REGION Network 7 (SCL): Head #4
   "M256_Manag_IDB".M256F_IDB[3].INPUT_xPressureDec :="i.1B414AP1.1B414SA1.Head4.CuttingPressure-";
   "M256_Manag_IDB".M256A_IDB[3].INPUT_xCarriageInWorkPosition := "i.1B414AP1.1B414SQ1.Head4.CarriageHeadWorkPosition";
   "M256_Manag_IDB".M256F_IDB[3].INPUT_xPressureInc := "i.1B414AP1.1B414SA1.Head4.CuttingPressure+";
   "Z256".INPUT_rgxHeadsInProduction[3] := "i.1B414AP1.1B414SA2.Head4.ProductionON";
   "M256_Manag_IDB".M256F_IDB[3].INPUT_xForceFiring := 0;
   "M256_Manag_IDB".M256A_IDB[3].INPUT_xForceArming := 0;
   "M256_Manag_IDB".M256M_IDB[3].INPUT_xBrakeRelease := FALSE;
   "M256_Manag_IDB".M256M_IDB[3].INPUT_xOverstroke := TRUE;//"i.1B410AP1.1B291KA4.Head4-5.CarriageTraslationAntiCollision";
END_REGION

REGION Network 8 (SCL): Head #5
   "M256_Manag_IDB".M256F_IDB[4].INPUT_xPressureDec := "i.1B415AP1.1B415SA1.Head5.CuttingPressure-";
   "M256_Manag_IDB".M256A_IDB[4].INPUT_xCarriageInWorkPosition := "i.1B415AP1.1B415SQ1.Head5.CarriageHeadWorkPosition";
   "M256_Manag_IDB".M256F_IDB[4].INPUT_xPressureInc := "i.1B415AP1.1B415SA1.Head5.CuttingPressure+";
   "Z256".INPUT_rgxHeadsInProduction[4] :="i.1B415AP1.1B415SA2.Head5.ProductionON";
   "M256_Manag_IDB".M256F_IDB[4].INPUT_xForceFiring := 0;
   "M256_Manag_IDB".M256A_IDB[4].INPUT_xForceArming := 0;
   "M256_Manag_IDB".M256M_IDB[4].INPUT_xBrakeRelease := FALSE;
   "M256_Manag_IDB".M256M_IDB[4].INPUT_xOverstroke := TRUE;//"i.1B410AP1.1B291KA5.Head5-6.CarriageTraslationAntiCollision";
END_REGION

REGION Network 9 (SCL): Head #6 / Head #5
   "M256_Manag_IDB".M256F_IDB[5].INPUT_xPressureDec := "i.1B416AP1.1B416SA1.Head6.CuttingPressure-";
   "M256_Manag_IDB".M256A_IDB[5].INPUT_xCarriageInWorkPosition := "i.1B416AP1.1B416SQ1.Head6.CarriageHeadWorkPosition";
   "M256_Manag_IDB".M256F_IDB[5].INPUT_xPressureInc := "i.1B416AP1.1B416SA1.Head6.CuttingPressure+";
   "Z256".INPUT_rgxHeadsInProduction[5] :="i.1B416AP1.1B416SA2.Head6.ProductionON";
   "M256_Manag_IDB".M256F_IDB[5].INPUT_xForceFiring := 0;
   "M256_Manag_IDB".M256A_IDB[5].INPUT_xForceArming := 0;
   "M256_Manag_IDB".M256M_IDB[5].INPUT_xBrakeRelease := FALSE;
   "M256_Manag_IDB".M256M_IDB[5].INPUT_xOverstroke := TRUE;//"i.1B410AP1.1B291KA8.Head6-7.CarriageTraslationAntiCollision";
END_REGION

REGION Network 10 (SCL): Head #7 / Head #5
   "M256_Manag_IDB".M256F_IDB[6].INPUT_xPressureDec := "i.1B417AP1.1B417SA1.Head7.CuttingPressure-";
   "M256_Manag_IDB".M256A_IDB[6].INPUT_xCarriageInWorkPosition := "i.1B417AP1.1B417SQ1.Head7.CarriageHeadWorkPosition";
   "M256_Manag_IDB".M256F_IDB[6].INPUT_xPressureInc := "i.1B417AP1.1B417SA1.Head7.CuttingPressure+";
   "Z256".INPUT_rgxHeadsInProduction[6] :="i.1B417AP1.1B417SA2.Head7.ProductionON";
   "M256_Manag_IDB".M256F_IDB[6].INPUT_xForceFiring := 0;
   "M256_Manag_IDB".M256A_IDB[6].INPUT_xForceArming := 0;
   "M256_Manag_IDB".M256M_IDB[6].INPUT_xBrakeRelease := FALSE;
   "M256_Manag_IDB".M256M_IDB[6].INPUT_xOverstroke := TRUE;//"i.1B410AP1.1B291KA7.Head7-8.CarriageTraslationAntiCollision";
END_REGION

REGION Network 11 (SCL): Head #8 / Head #5
   "M256_Manag_IDB".M256F_IDB[7].INPUT_xPressureDec := "i.1B418AP1.1B418SA1.Head8.CuttingPressure-";
   "M256_Manag_IDB".M256A_IDB[7].INPUT_xCarriageInWorkPosition := "i.1B418AP1.1B418SQ1.Head8.CarriageHeadWorkPosition";
   "M256_Manag_IDB".M256F_IDB[7].INPUT_xPressureInc := "i.1B418AP1.1B418SA1.Head8.CuttingPressure+";
   "Z256".INPUT_rgxHeadsInProduction[7] :="i.1B418AP1.1B418SA2.Head8.ProductionON";
   "M256_Manag_IDB".M256F_IDB[7].INPUT_xForceFiring := 0;
   "M256_Manag_IDB".M256A_IDB[7].INPUT_xForceArming := 0;
   "M256_Manag_IDB".M256M_IDB[7].INPUT_xBrakeRelease := FALSE;
   "M256_Manag_IDB".M256M_IDB[7].INPUT_xOverstroke := TRUE;//"i.1B410AP1.1B291KA8.Head8-9.CarriageTraslationAntiCollision";
END_REGION

REGION Network 12 (SCL): IDevice
   "CM_IDEV_FromMainLine" := "i.IDeviceCPU0";
END_REGION
END_FUNCTION

FUNCTION "M256M_SbrCheckCollision" : Void   // FC10, SCL
{ S7_Optimized_Access := 'TRUE' }
VERSION : 0.1
   VAR_OUTPUT
      o_rgxHeadVirtualCollision : Array[0.."CONST_dNumberOfHeadsCycle"] of Bool;
   END_VAR
   VAR_TEMP
      TMP_dIndex : DInt;
      TMP_xCollision : Bool;
      TMP_xCollisionNext : Bool;
      TMP_dActHeadPosition_cmm : DInt;
      TMP_dNextHeadPosition_cmm : DInt;
   END_VAR
BEGIN
   ////--------------------------------------------------------------------------------------------------------------------
   //   Copyright (c)  Bottero Spa
   //--------------------------------------------------------------
   //   Routine: NomeRoutine
   //       Author: Alberto Cigliutti
   //   Created: July 2016
   //--------------------------------------------------------------
   //   Description: This routine will analize the data out from the manager, and compile 
   //  a collision array
   //
   //   History:
   //
   ////--------------------------------------------------------------------------------------------------------------------

   FOR #TMP_dIndex := 0 TO "CONST_dNumberOfHeadsCycle" DO
       #o_rgxHeadVirtualCollision[#TMP_dIndex] := 0;
   END_FOR;

   FOR #TMP_dIndex := 0 TO "CONST_dNumberOfHeadsCycle" DO

       #TMP_xCollision := 0;
       #TMP_xCollisionNext := 0;

       IF #TMP_dIndex = 0 OR #TMP_dIndex = "CONST_dNumberOfHeadsCycle" THEN
           //For the first head and last head, we check the position request, if is less then the home
           //we rise a virtual collision
           IF NOT "PLANT_CONSTANTS".CONST_rgxHomeSide[#TMP_dIndex] AND
               ("Z256_Manager".tOutputData.rgdHeadsPositions_cmm[#TMP_dIndex] < "M256_Manag_IDB".M256M_IDB[#TMP_dIndex].tHMR.dHeadHomePositions_cmm) THEN

               #TMP_xCollision := 1;
               #o_rgxHeadVirtualCollision[#TMP_dIndex] := #TMP_xCollision;

           ELSIF ("PLANT_CONSTANTS".CONST_rgxHomeSide[#TMP_dIndex] AND
               "Z256_Manager".tOutputData.rgdHeadsPositions_cmm[#TMP_dIndex]>"M256_Manag_IDB".M256M_IDB[#TMP_dIndex].tHMR.dHeadHomePositions_cmm) THEN

               #TMP_xCollision := 1;
               #o_rgxHeadVirtualCollision[#TMP_dIndex] := #TMP_xCollision;
           END_IF;
       END_IF;

       //Start to search the next head position,
       //only jump this check on the last head
       IF #TMP_dIndex < "CONST_dNumberOfHeadsCycle" THEN

           #TMP_dActHeadPosition_cmm := "Z256_Manager".tOutputData.rgdHeadsPositions_cmm[#TMP_dIndex] + "PLANT_CONSTANTS".CONST_dHOppoSideEnc_cmm[#TMP_dIndex];
           #TMP_dNextHeadPosition_cmm := "Z256_Manager".tOutputData.rgdHeadsPositions_cmm[#TMP_dIndex + 1] - "PLANT_CONSTANTS".CONST_dHOpSideEnc_cmm[#TMP_dIndex + 1];

           IF (#TMP_dActHeadPosition_cmm > #TMP_dNextHeadPosition_cmm) THEN
               #TMP_xCollision := 1;
               #TMP_xCollisionNext := 1;
           END_IF;

           #o_rgxHeadVirtualCollision[#TMP_dIndex + 1] := #TMP_xCollisionNext;
           #o_rgxHeadVirtualCollision[#TMP_dIndex] := #TMP_xCollision;

       END_IF;



   END_FOR;
END_FUNCTION

FUNCTION "M256M_HMI_Logics" : Void   // FC11, LAD
{ S7_Optimized_Access := 'TRUE' }
VERSION : 0.1
   VAR_IN_OUT
      io_ST_xHeadReferredSwitch : Array[0.."CONST_dNumberOfHeadsCycle"] of Bool;
   END_VAR
   VAR_TEMP
      TMP_dIndex : DInt;
   END_VAR
   VAR_TEMP   // added for the SCL form of the ladder/FBD networks
      _w1 : Bool;
   END_VAR
BEGIN

REGION Network 1: #####_HMI_LOGICS_#####
END_REGION

REGION Network 2 (SCL): Force heads homing
   IF "Z256_hmi".tHMW.xForceHeadsHoming THEN
       FOR #TMP_dIndex := 0 TO "CONST_dNumberOfHeadsCycle" DO
           #io_ST_xHeadReferredSwitch[#TMP_dIndex] := 0;
       END_FOR;
       "Z256_hmi".tHMW.xForceHeadsHoming := false;
   END_IF;
END_REGION

REGION Network 3: Calibration function allowed
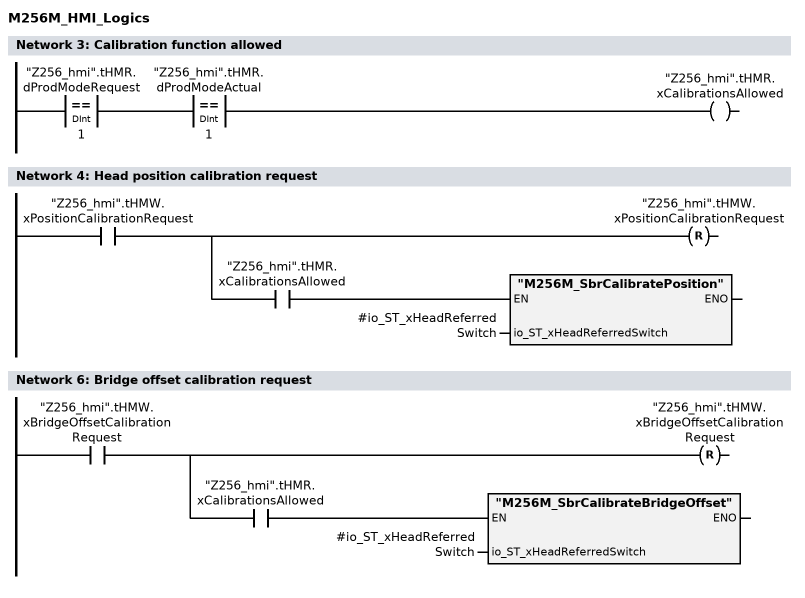
   RUNG wire#powerrail
      { S7_Templates := "SrcType := DInt" } EQ_Contact(in1 := "Z256_hmi".tHMR.dProdModeRequest, in2 := 1)
      { S7_Templates := "SrcType := DInt" } EQ_Contact(in1 := "Z256_hmi".tHMR.dProdModeActual, in2 := 1)
      Coil( "Z256_hmi".tHMR.xCalibrationsAllowed )
   END_RUNG
   // the same network as SCL:
   "Z256_hmi".tHMR.xCalibrationsAllowed := ("Z256_hmi".tHMR.dProdModeRequest = 1) AND ("Z256_hmi".tHMR.dProdModeActual = 1);
END_REGION

REGION Network 4: Head position calibration request
   RUNG wire#powerrail
      Contact( "Z256_hmi".tHMW.xPositionCalibrationRequest )
      wire#w1
      R_Coil( "Z256_hmi".tHMW.xPositionCalibrationRequest )
   END_RUNG
   RUNG wire#w1
      Contact( "Z256_hmi".tHMR.xCalibrationsAllowed )
      "M256M_SbrCalibratePosition"(io_ST_xHeadReferredSwitch := #io_ST_xHeadReferredSwitch)
   END_RUNG
   // the same network as SCL:
   #_w1 := "Z256_hmi".tHMW.xPositionCalibrationRequest;
   IF #_w1 THEN "Z256_hmi".tHMW.xPositionCalibrationRequest := FALSE; END_IF;
   IF #_w1 AND "Z256_hmi".tHMR.xCalibrationsAllowed THEN
       "M256M_SbrCalibratePosition"(io_ST_xHeadReferredSwitch := #io_ST_xHeadReferredSwitch);
   END_IF;
END_REGION

REGION Network 5 (SCL): Update home head
   FOR #TMP_dIndex := 0 TO "CONST_dNumberOfHeadsCycle" DO
       IF "M256_Manag_IDB".M256M_IDB[#TMP_dIndex].tHMW.xUpdateHomeHead THEN
           "M256_Manag_IDB".M256M_IDB[#TMP_dIndex].tHMW.xUpdateHomeHead := 0; 
           "M256_Manag_IDB".M256M_IDB[#TMP_dIndex].tHMR.dHeadHomePositions_cmm := "M256_Manag_IDB".M256M_IDB[#TMP_dIndex].tHMW.dHeadHomePositions_cmm;
       END_IF;
   END_FOR;
END_REGION

REGION Network 6: Bridge offset calibration request
   RUNG wire#powerrail
      Contact( "Z256_hmi".tHMW.xBridgeOffsetCalibrationRequest )
      wire#w1
      R_Coil( "Z256_hmi".tHMW.xBridgeOffsetCalibrationRequest )
   END_RUNG
   RUNG wire#w1
      Contact( "Z256_hmi".tHMR.xCalibrationsAllowed )
      "M256M_SbrCalibrateBridgeOffset"(io_ST_xHeadReferredSwitch := #io_ST_xHeadReferredSwitch)
   END_RUNG
   // the same network as SCL:
   #_w1 := "Z256_hmi".tHMW.xBridgeOffsetCalibrationRequest;
   IF #_w1 THEN "Z256_hmi".tHMW.xBridgeOffsetCalibrationRequest := FALSE; END_IF;
   IF #_w1 AND "Z256_hmi".tHMR.xCalibrationsAllowed THEN
       "M256M_SbrCalibrateBridgeOffset"(io_ST_xHeadReferredSwitch := #io_ST_xHeadReferredSwitch);
   END_IF;
END_REGION
END_FUNCTION

FUNCTION "Encoder_Manager" : Void   // FC12, LAD
{ S7_Optimized_Access := 'TRUE' }
VERSION : 0.1
   VAR_TEMP
      TMP_rDummy : Real;
      TMP_dDummy : DInt;
      TMP_dIndex : DInt;
   END_VAR
   VAR_TEMP   // added for the SCL form of the ladder/FBD networks
      _w1 : Bool;
   END_VAR
BEGIN

REGION Network 1: Enable card counter
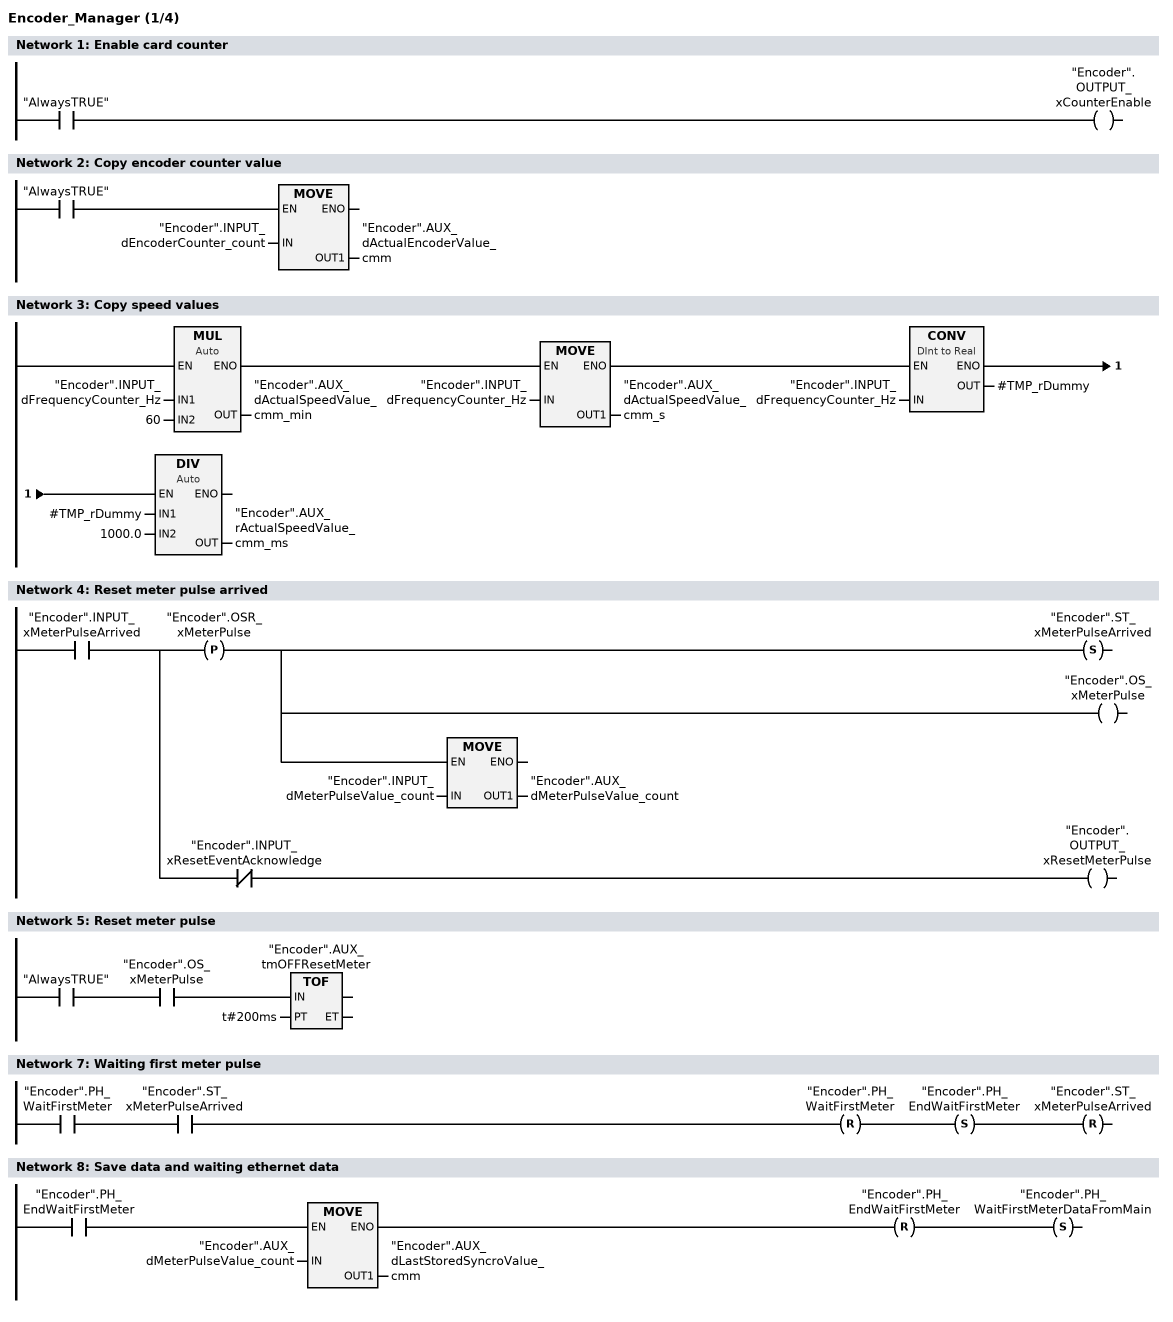
   RUNG wire#powerrail
      Contact( "AlwaysTRUE" )
      Coil( "Encoder".OUTPUT_xCounterEnable )
   END_RUNG
   // the same network as SCL:
   "Encoder".OUTPUT_xCounterEnable := "AlwaysTRUE";
END_REGION

REGION Network 2: Copy encoder counter value
   RUNG wire#powerrail
      Contact( "AlwaysTRUE" )
      Move(in := "Encoder".INPUT_dEncoderCounter_count, out1 => "Encoder".AUX_dActualEncoderValue_cmm)
   END_RUNG
   // the same network as SCL:
   IF "AlwaysTRUE" THEN
       "Encoder".AUX_dActualEncoderValue_cmm := "Encoder".INPUT_dEncoderCounter_count;
   END_IF;
END_REGION

REGION Network 3: Copy speed values
   RUNG wire#powerrail
      Mul(in1 := "Encoder".INPUT_dFrequencyCounter_Hz, in2 := 60, out => "Encoder".AUX_dActualSpeedValue_cmm_min)
      Move(in := "Encoder".INPUT_dFrequencyCounter_Hz, out1 => "Encoder".AUX_dActualSpeedValue_cmm_s)
      { S7_Templates := "[SrcType := DInt, DestType := Real]" } Convert(in := "Encoder".INPUT_dFrequencyCounter_Hz, out => #TMP_rDummy)
      Div(in1 := #TMP_rDummy, in2 := 1000.0, out => "Encoder".AUX_rActualSpeedValue_cmm_ms)
   END_RUNG
   // the same network as SCL:
   "Encoder".AUX_dActualSpeedValue_cmm_min := "Encoder".INPUT_dFrequencyCounter_Hz * 60;
   "Encoder".AUX_dActualSpeedValue_cmm_s := "Encoder".INPUT_dFrequencyCounter_Hz;
   #TMP_rDummy := DINT_TO_REAL("Encoder".INPUT_dFrequencyCounter_Hz);
   "Encoder".AUX_rActualSpeedValue_cmm_ms := #TMP_rDummy / 1000.0;
END_REGION

REGION Network 4: Reset meter pulse arrived
   RUNG wire#powerrail
      Contact( "Encoder".INPUT_xMeterPulseArrived )
      wire#w1
      P_Trig( "Encoder".OSR_xMeterPulse )
      wire#w2
      S_Coil( "Encoder".ST_xMeterPulseArrived )
   END_RUNG
   RUNG wire#w2
      Coil( "Encoder".OS_xMeterPulse )
   END_RUNG
   RUNG wire#w2
      Move(in := "Encoder".INPUT_dMeterPulseValue_count, out1 => "Encoder".AUX_dMeterPulseValue_count)
   END_RUNG
   RUNG wire#w1
      I_Contact( "Encoder".INPUT_xResetEventAcknowledge )
      Coil( "Encoder".OUTPUT_xResetMeterPulse )
   END_RUNG
   // the same network as SCL:
   #_w1 := "Encoder".INPUT_xMeterPulseArrived AND NOT "Encoder".OSR_xMeterPulse;   // rising edge
   "Encoder".OSR_xMeterPulse := "Encoder".INPUT_xMeterPulseArrived;
   IF #_w1 THEN "Encoder".ST_xMeterPulseArrived := TRUE; END_IF;
   "Encoder".OS_xMeterPulse := #_w1;
   IF #_w1 THEN "Encoder".AUX_dMeterPulseValue_count := "Encoder".INPUT_dMeterPulseValue_count; END_IF;
   "Encoder".OUTPUT_xResetMeterPulse := "Encoder".INPUT_xMeterPulseArrived AND NOT "Encoder".INPUT_xResetEventAcknowledge;
END_REGION

REGION Network 5: Reset meter pulse
   "Encoder".AUX_tmOFFResetMeter.TOF(IN := "AlwaysTRUE" AND "Encoder".OS_xMeterPulse, PT := t#200ms);
END_REGION

REGION Network 6: ### FIRST METER PHASES ###
END_REGION

REGION Network 7: Waiting first meter pulse
   RUNG wire#powerrail
      Contact( "Encoder".PH_WaitFirstMeter )
      Contact( "Encoder".ST_xMeterPulseArrived )
      R_Coil( "Encoder".PH_WaitFirstMeter )
      S_Coil( "Encoder".PH_EndWaitFirstMeter )
      R_Coil( "Encoder".ST_xMeterPulseArrived )
   END_RUNG
   // the same network as SCL:
   #_w1 := "Encoder".PH_WaitFirstMeter AND "Encoder".ST_xMeterPulseArrived;
   IF #_w1 THEN
       "Encoder".PH_WaitFirstMeter := FALSE;
       "Encoder".PH_EndWaitFirstMeter := TRUE;
       "Encoder".ST_xMeterPulseArrived := FALSE;
   END_IF;
END_REGION

REGION Network 8: Save data and waiting ethernet data
   RUNG wire#powerrail
      Contact( "Encoder".PH_EndWaitFirstMeter )
      Move(in := "Encoder".AUX_dMeterPulseValue_count, out1 => "Encoder".AUX_dLastStoredSyncroValue_cmm)
      R_Coil( "Encoder".PH_EndWaitFirstMeter )
      S_Coil( "Encoder".PH_WaitFirstMeterDataFromMain )
   END_RUNG
   // the same network as SCL:
   IF "Encoder".PH_EndWaitFirstMeter THEN
       "Encoder".AUX_dLastStoredSyncroValue_cmm := "Encoder".AUX_dMeterPulseValue_count;
   END_IF;
   #_w1 := "Encoder".PH_EndWaitFirstMeter;
   IF #_w1 THEN
       "Encoder".PH_EndWaitFirstMeter := FALSE;
       "Encoder".PH_WaitFirstMeterDataFromMain := TRUE;
   END_IF;
END_REGION

REGION Network 9: End waiting ethernet data
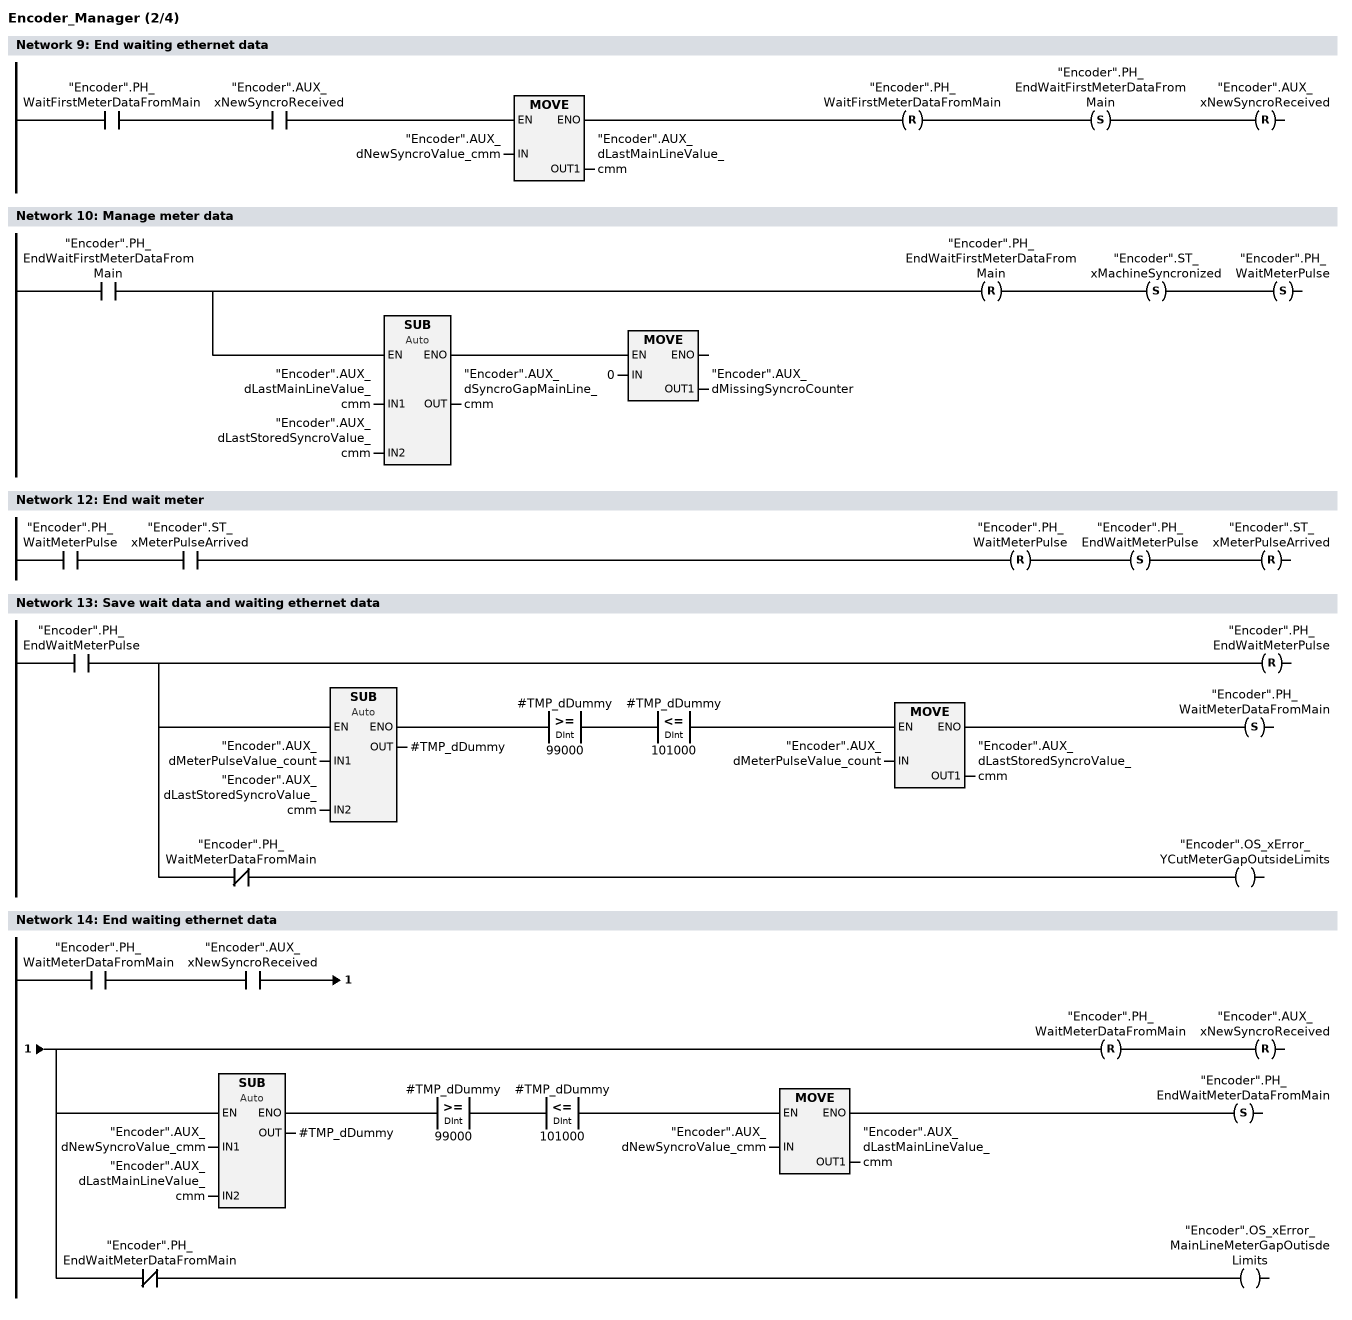
   RUNG wire#powerrail
      Contact( "Encoder".PH_WaitFirstMeterDataFromMain )
      Contact( "Encoder".AUX_xNewSyncroReceived )
      Move(in := "Encoder".AUX_dNewSyncroValue_cmm, out1 => "Encoder".AUX_dLastMainLineValue_cmm)
      R_Coil( "Encoder".PH_WaitFirstMeterDataFromMain )
      S_Coil( "Encoder".PH_EndWaitFirstMeterDataFromMain )
      R_Coil( "Encoder".AUX_xNewSyncroReceived )
   END_RUNG
   // the same network as SCL:
   IF "Encoder".PH_WaitFirstMeterDataFromMain AND "Encoder".AUX_xNewSyncroReceived THEN
       "Encoder".AUX_dLastMainLineValue_cmm := "Encoder".AUX_dNewSyncroValue_cmm;
   END_IF;
   #_w1 := "Encoder".PH_WaitFirstMeterDataFromMain AND "Encoder".AUX_xNewSyncroReceived;
   IF #_w1 THEN
       "Encoder".PH_WaitFirstMeterDataFromMain := FALSE;
       "Encoder".PH_EndWaitFirstMeterDataFromMain := TRUE;
       "Encoder".AUX_xNewSyncroReceived := FALSE;
   END_IF;
END_REGION

REGION Network 10: Manage meter data
   RUNG wire#powerrail
      Contact( "Encoder".PH_EndWaitFirstMeterDataFromMain )
      wire#w1
      R_Coil( "Encoder".PH_EndWaitFirstMeterDataFromMain )
      S_Coil( "Encoder".ST_xMachineSyncronized )
      S_Coil( "Encoder".PH_WaitMeterPulse )
   END_RUNG
   RUNG wire#w1
      Sub(in1 := "Encoder".AUX_dLastMainLineValue_cmm, in2 := "Encoder".AUX_dLastStoredSyncroValue_cmm, out => "Encoder".AUX_dSyncroGapMainLine_cmm)
      Move(in := 0, out1 => "Encoder".AUX_dMissingSyncroCounter)
   END_RUNG
   // the same network as SCL:
   #_w1 := "Encoder".PH_EndWaitFirstMeterDataFromMain;
   IF #_w1 THEN
       "Encoder".PH_EndWaitFirstMeterDataFromMain := FALSE;
       "Encoder".ST_xMachineSyncronized := TRUE;
       "Encoder".PH_WaitMeterPulse := TRUE;
       "Encoder".AUX_dSyncroGapMainLine_cmm := "Encoder".AUX_dLastMainLineValue_cmm - "Encoder".AUX_dLastStoredSyncroValue_cmm;
       "Encoder".AUX_dMissingSyncroCounter := 0;
   END_IF;
END_REGION

REGION Network 11: ### METER PHASES ###
END_REGION

REGION Network 12: End wait meter
   RUNG wire#powerrail
      Contact( "Encoder".PH_WaitMeterPulse )
      Contact( "Encoder".ST_xMeterPulseArrived )
      R_Coil( "Encoder".PH_WaitMeterPulse )
      S_Coil( "Encoder".PH_EndWaitMeterPulse )
      R_Coil( "Encoder".ST_xMeterPulseArrived )
   END_RUNG
   // the same network as SCL:
   #_w1 := "Encoder".PH_WaitMeterPulse AND "Encoder".ST_xMeterPulseArrived;
   IF #_w1 THEN
       "Encoder".PH_WaitMeterPulse := FALSE;
       "Encoder".PH_EndWaitMeterPulse := TRUE;
       "Encoder".ST_xMeterPulseArrived := FALSE;
   END_IF;
END_REGION

REGION Network 13: Save wait data and waiting ethernet data
   RUNG wire#powerrail
      Contact( "Encoder".PH_EndWaitMeterPulse )
      wire#w1
      R_Coil( "Encoder".PH_EndWaitMeterPulse )
   END_RUNG
   RUNG wire#w1
      Sub(in1 := "Encoder".AUX_dMeterPulseValue_count, in2 := "Encoder".AUX_dLastStoredSyncroValue_cmm, out => #TMP_dDummy)
      { S7_Templates := "SrcType := DInt" } GE_Contact(in1 := #TMP_dDummy, in2 := 99000)
      { S7_Templates := "SrcType := DInt" } LE_Contact(in1 := #TMP_dDummy, in2 := 101000)
      Move(in := "Encoder".AUX_dMeterPulseValue_count, out1 => "Encoder".AUX_dLastStoredSyncroValue_cmm)
      S_Coil( "Encoder".PH_WaitMeterDataFromMain )
   END_RUNG
   RUNG wire#w1
      I_Contact( "Encoder".PH_WaitMeterDataFromMain )
      Coil( "Encoder".OS_xError_YCutMeterGapOutsideLimits )
   END_RUNG
   // the same network as SCL:
   #_w1 := "Encoder".PH_EndWaitMeterPulse;
   IF #_w1 THEN
       "Encoder".PH_EndWaitMeterPulse := FALSE;
       #TMP_dDummy := "Encoder".AUX_dMeterPulseValue_count - "Encoder".AUX_dLastStoredSyncroValue_cmm;
   END_IF;
   IF #_w1 AND (#TMP_dDummy >= 99000) AND (#TMP_dDummy <= 101000) THEN
       "Encoder".AUX_dLastStoredSyncroValue_cmm := "Encoder".AUX_dMeterPulseValue_count;
       "Encoder".PH_WaitMeterDataFromMain := TRUE;
   END_IF;
   "Encoder".OS_xError_YCutMeterGapOutsideLimits := #_w1 AND NOT "Encoder".PH_WaitMeterDataFromMain;
END_REGION

REGION Network 14: End waiting ethernet data
   RUNG wire#powerrail
      Contact( "Encoder".PH_WaitMeterDataFromMain )
      Contact( "Encoder".AUX_xNewSyncroReceived )
      wire#w1
      R_Coil( "Encoder".PH_WaitMeterDataFromMain )
      R_Coil( "Encoder".AUX_xNewSyncroReceived )
   END_RUNG
   RUNG wire#w1
      Sub(in1 := "Encoder".AUX_dNewSyncroValue_cmm, in2 := "Encoder".AUX_dLastMainLineValue_cmm, out => #TMP_dDummy)
      { S7_Templates := "SrcType := DInt" } GE_Contact(in1 := #TMP_dDummy, in2 := 99000)
      { S7_Templates := "SrcType := DInt" } LE_Contact(in1 := #TMP_dDummy, in2 := 101000)
      Move(in := "Encoder".AUX_dNewSyncroValue_cmm, out1 => "Encoder".AUX_dLastMainLineValue_cmm)
      S_Coil( "Encoder".PH_EndWaitMeterDataFromMain )
   END_RUNG
   RUNG wire#w1
      I_Contact( "Encoder".PH_EndWaitMeterDataFromMain )
      Coil( "Encoder".OS_xError_MainLineMeterGapOutisdeLimits )
   END_RUNG
   // the same network as SCL:
   #_w1 := "Encoder".PH_WaitMeterDataFromMain AND "Encoder".AUX_xNewSyncroReceived;
   IF #_w1 THEN
       "Encoder".PH_WaitMeterDataFromMain := FALSE;
       "Encoder".AUX_xNewSyncroReceived := FALSE;
       #TMP_dDummy := "Encoder".AUX_dNewSyncroValue_cmm - "Encoder".AUX_dLastMainLineValue_cmm;
   END_IF;
   IF #_w1 AND (#TMP_dDummy >= 99000) AND (#TMP_dDummy <= 101000) THEN
       "Encoder".AUX_dLastMainLineValue_cmm := "Encoder".AUX_dNewSyncroValue_cmm;
       "Encoder".PH_EndWaitMeterDataFromMain := TRUE;
   END_IF;
   "Encoder".OS_xError_MainLineMeterGapOutisdeLimits := #_w1 AND NOT "Encoder".PH_EndWaitMeterDataFromMain;
END_REGION

REGION Network 15: Manage meter data
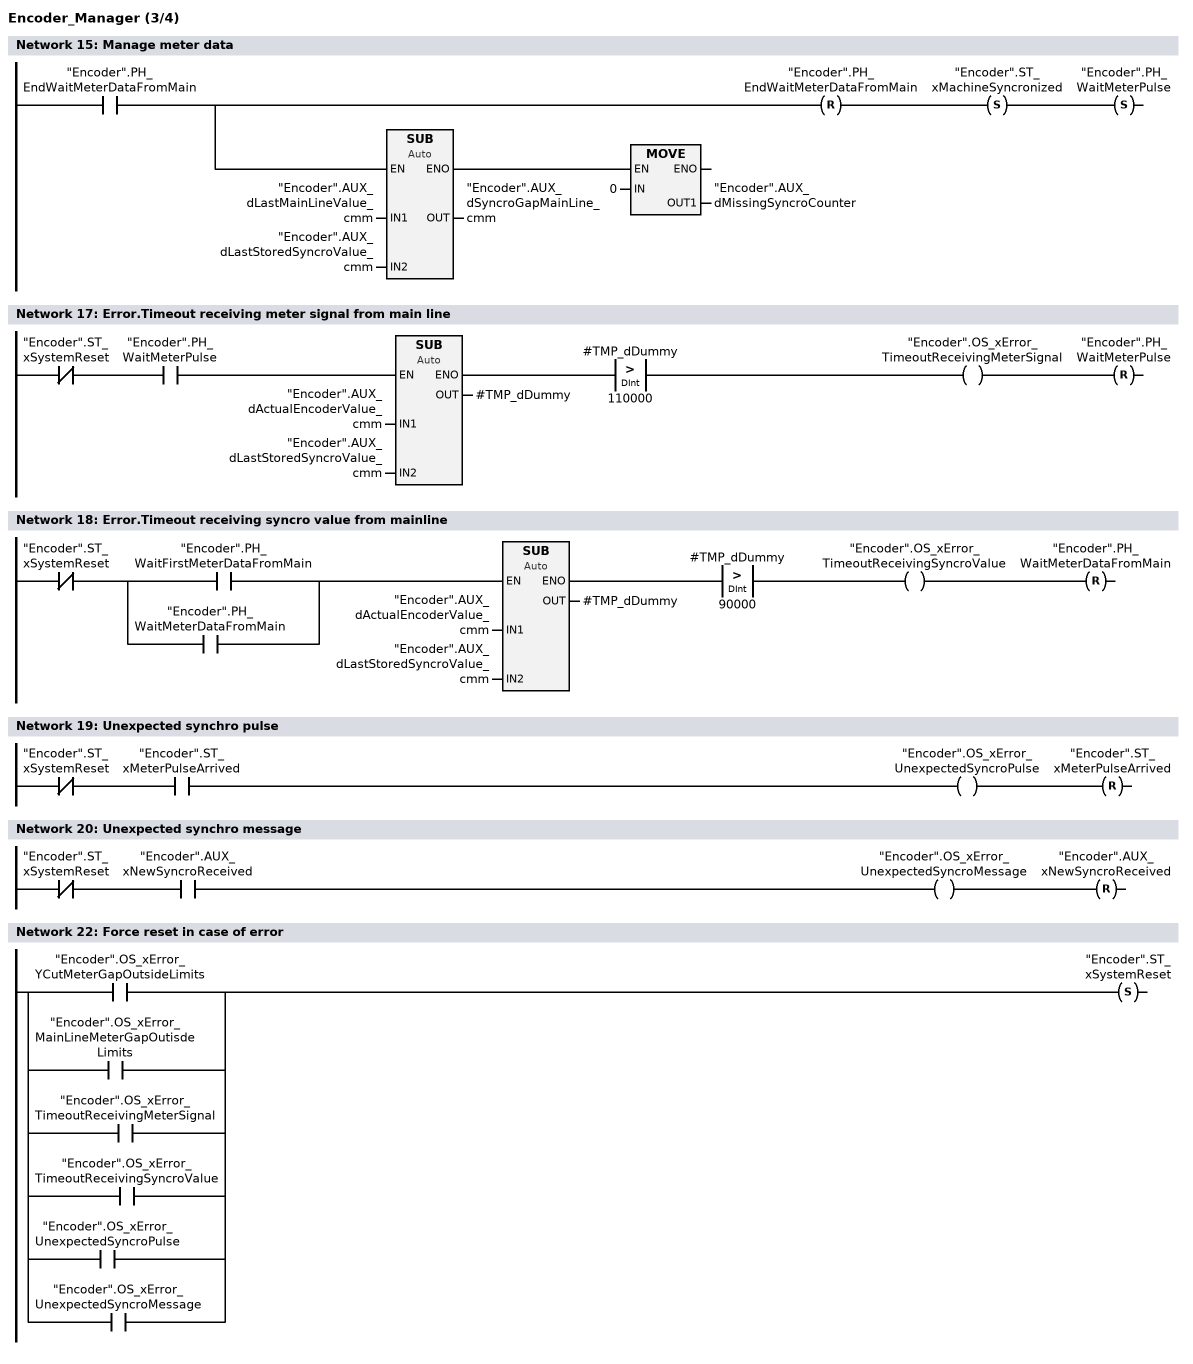
   RUNG wire#powerrail
      Contact( "Encoder".PH_EndWaitMeterDataFromMain )
      wire#w1
      R_Coil( "Encoder".PH_EndWaitMeterDataFromMain )
      S_Coil( "Encoder".ST_xMachineSyncronized )
      S_Coil( "Encoder".PH_WaitMeterPulse )
   END_RUNG
   RUNG wire#w1
      Sub(in1 := "Encoder".AUX_dLastMainLineValue_cmm, in2 := "Encoder".AUX_dLastStoredSyncroValue_cmm, out => "Encoder".AUX_dSyncroGapMainLine_cmm)
      Move(in := 0, out1 => "Encoder".AUX_dMissingSyncroCounter)
   END_RUNG
   // the same network as SCL:
   #_w1 := "Encoder".PH_EndWaitMeterDataFromMain;
   IF #_w1 THEN
       "Encoder".PH_EndWaitMeterDataFromMain := FALSE;
       "Encoder".ST_xMachineSyncronized := TRUE;
       "Encoder".PH_WaitMeterPulse := TRUE;
       "Encoder".AUX_dSyncroGapMainLine_cmm := "Encoder".AUX_dLastMainLineValue_cmm - "Encoder".AUX_dLastStoredSyncroValue_cmm;
       "Encoder".AUX_dMissingSyncroCounter := 0;
   END_IF;
END_REGION

REGION Network 16: ### ERRORS AND TIMEOUTS ###
END_REGION

REGION Network 17: Error.Timeout receiving meter signal from main line
   RUNG wire#powerrail
      I_Contact( "Encoder".ST_xSystemReset )
      Contact( "Encoder".PH_WaitMeterPulse )
      Sub(in1 := "Encoder".AUX_dActualEncoderValue_cmm, in2 := "Encoder".AUX_dLastStoredSyncroValue_cmm, out => #TMP_dDummy)
      { S7_Templates := "SrcType := DInt" } GT_Contact(in1 := #TMP_dDummy, in2 := 110000)
      Coil( "Encoder".OS_xError_TimeoutReceivingMeterSignal )
      R_Coil( "Encoder".PH_WaitMeterPulse )
   END_RUNG
   // the same network as SCL:
   #_w1 := NOT "Encoder".ST_xSystemReset AND "Encoder".PH_WaitMeterPulse;
   IF #_w1 THEN
       #TMP_dDummy := "Encoder".AUX_dActualEncoderValue_cmm - "Encoder".AUX_dLastStoredSyncroValue_cmm;
   END_IF;
   "Encoder".OS_xError_TimeoutReceivingMeterSignal := #_w1 AND (#TMP_dDummy > 110000);
   IF "Encoder".OS_xError_TimeoutReceivingMeterSignal THEN "Encoder".PH_WaitMeterPulse := FALSE; END_IF;
END_REGION

REGION Network 18: Error.Timeout receiving syncro value from mainline
   RUNG wire#powerrail
      I_Contact( "Encoder".ST_xSystemReset )
      wire#w1
      Contact( "Encoder".PH_WaitFirstMeterDataFromMain )
      wire#w2
      Sub(in1 := "Encoder".AUX_dActualEncoderValue_cmm, in2 := "Encoder".AUX_dLastStoredSyncroValue_cmm, out => #TMP_dDummy)
      { S7_Templates := "SrcType := DInt" } GT_Contact(in1 := #TMP_dDummy, in2 := 90000)
      Coil( "Encoder".OS_xError_TimeoutReceivingSyncroValue )
      R_Coil( "Encoder".PH_WaitMeterDataFromMain )
   END_RUNG
   RUNG wire#w1
      Contact( "Encoder".PH_WaitMeterDataFromMain )
   END_RUNG wire#w2
   // the same network as SCL:
   #_w1 := NOT "Encoder".ST_xSystemReset AND ("Encoder".PH_WaitFirstMeterDataFromMain OR "Encoder".PH_WaitMeterDataFromMain);
   IF #_w1 THEN
       #TMP_dDummy := "Encoder".AUX_dActualEncoderValue_cmm - "Encoder".AUX_dLastStoredSyncroValue_cmm;
   END_IF;
   "Encoder".OS_xError_TimeoutReceivingSyncroValue := #_w1 AND (#TMP_dDummy > 90000);
   IF "Encoder".OS_xError_TimeoutReceivingSyncroValue THEN
       "Encoder".PH_WaitMeterDataFromMain := FALSE;
   END_IF;
END_REGION

REGION Network 19: Unexpected synchro pulse
   RUNG wire#powerrail
      I_Contact( "Encoder".ST_xSystemReset )
      Contact( "Encoder".ST_xMeterPulseArrived )
      Coil( "Encoder".OS_xError_UnexpectedSyncroPulse )
      R_Coil( "Encoder".ST_xMeterPulseArrived )
   END_RUNG
   // the same network as SCL:
   "Encoder".OS_xError_UnexpectedSyncroPulse := NOT "Encoder".ST_xSystemReset AND "Encoder".ST_xMeterPulseArrived;
   IF "Encoder".OS_xError_UnexpectedSyncroPulse THEN "Encoder".ST_xMeterPulseArrived := FALSE; END_IF;
END_REGION

REGION Network 20: Unexpected synchro message
   RUNG wire#powerrail
      I_Contact( "Encoder".ST_xSystemReset )
      Contact( "Encoder".AUX_xNewSyncroReceived )
      Coil( "Encoder".OS_xError_UnexpectedSyncroMessage )
      R_Coil( "Encoder".AUX_xNewSyncroReceived )
   END_RUNG
   // the same network as SCL:
   "Encoder".OS_xError_UnexpectedSyncroMessage := NOT "Encoder".ST_xSystemReset AND "Encoder".AUX_xNewSyncroReceived;
   IF "Encoder".OS_xError_UnexpectedSyncroMessage THEN "Encoder".AUX_xNewSyncroReceived := FALSE; END_IF;
END_REGION

REGION Network 21: ### RESET AND INITIALIZE CARD MANAGER ###
END_REGION

REGION Network 22: Force reset in case of error
   RUNG wire#powerrail
      Contact( "Encoder".OS_xError_YCutMeterGapOutsideLimits )
      wire#w1
      S_Coil( "Encoder".ST_xSystemReset )
   END_RUNG
   RUNG wire#powerrail
      Contact( "Encoder".OS_xError_MainLineMeterGapOutisdeLimits )
   END_RUNG wire#w1
   RUNG wire#powerrail
      Contact( "Encoder".OS_xError_TimeoutReceivingMeterSignal )
   END_RUNG wire#w1
   RUNG wire#powerrail
      Contact( "Encoder".OS_xError_TimeoutReceivingSyncroValue )
   END_RUNG wire#w1
   RUNG wire#powerrail
      Contact( "Encoder".OS_xError_UnexpectedSyncroPulse )
   END_RUNG wire#w1
   RUNG wire#powerrail
      Contact( "Encoder".OS_xError_UnexpectedSyncroMessage )
   END_RUNG wire#w1
   // the same network as SCL:
   IF "Encoder".OS_xError_YCutMeterGapOutsideLimits OR "Encoder".OS_xError_MainLineMeterGapOutisdeLimits OR "Encoder".OS_xError_TimeoutReceivingMeterSignal OR "Encoder".OS_xError_TimeoutReceivingSyncroValue OR "Encoder".OS_xError_UnexpectedSyncroPulse OR "Encoder".OS_xError_UnexpectedSyncroMessage THEN
       "Encoder".ST_xSystemReset := TRUE;
   END_IF;
END_REGION

REGION Network 23: Reset encoder counter
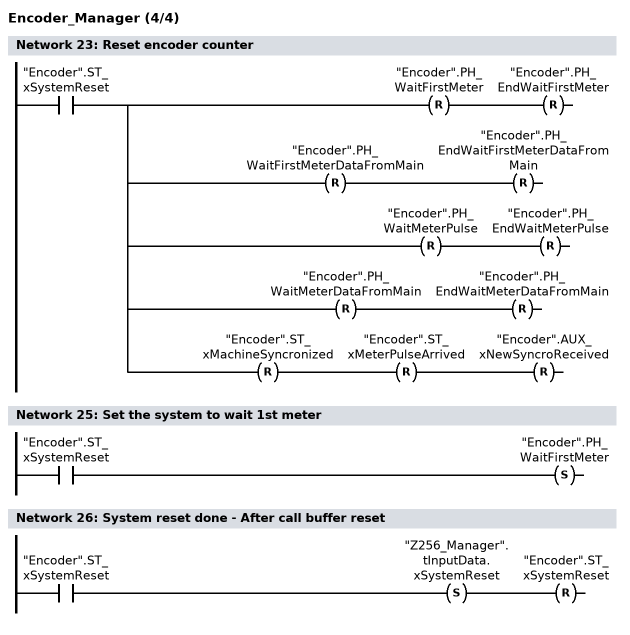
   RUNG wire#powerrail
      Contact( "Encoder".ST_xSystemReset )
      wire#w1
      R_Coil( "Encoder".PH_WaitFirstMeter )
      R_Coil( "Encoder".PH_EndWaitFirstMeter )
   END_RUNG
   RUNG wire#w1
      R_Coil( "Encoder".PH_WaitFirstMeterDataFromMain )
      R_Coil( "Encoder".PH_EndWaitFirstMeterDataFromMain )
   END_RUNG
   RUNG wire#w1
      R_Coil( "Encoder".PH_WaitMeterPulse )
      R_Coil( "Encoder".PH_EndWaitMeterPulse )
   END_RUNG
   RUNG wire#w1
      R_Coil( "Encoder".PH_WaitMeterDataFromMain )
      R_Coil( "Encoder".PH_EndWaitMeterDataFromMain )
   END_RUNG
   RUNG wire#w1
      R_Coil( "Encoder".ST_xMachineSyncronized )
      R_Coil( "Encoder".ST_xMeterPulseArrived )
      R_Coil( "Encoder".AUX_xNewSyncroReceived )
   END_RUNG
   // the same network as SCL:
   IF "Encoder".ST_xSystemReset THEN
       "Encoder".PH_WaitFirstMeter := FALSE;
       "Encoder".PH_EndWaitFirstMeter := FALSE;
       "Encoder".PH_WaitFirstMeterDataFromMain := FALSE;
       "Encoder".PH_EndWaitFirstMeterDataFromMain := FALSE;
       "Encoder".PH_WaitMeterPulse := FALSE;
       "Encoder".PH_EndWaitMeterPulse := FALSE;
       "Encoder".PH_WaitMeterDataFromMain := FALSE;
       "Encoder".PH_EndWaitMeterDataFromMain := FALSE;
       "Encoder".ST_xMachineSyncronized := FALSE;
       "Encoder".ST_xMeterPulseArrived := FALSE;
       "Encoder".AUX_xNewSyncroReceived := FALSE;
   END_IF;
END_REGION

REGION Network 24 (SCL): System reset
   IF "Encoder".ST_xSystemReset THEN
       FOR #TMP_dIndex := 0 TO "CONST_dNumberOfHeadsCycle" DO
           "M256_Manag_IDB".M256F_IDB[#TMP_dIndex].AUX_xHeadFiringMissionInProgress := 0;
       END_FOR;
   END_IF;
END_REGION

REGION Network 25: Set the system to wait 1st meter
   RUNG wire#powerrail
      Contact( "Encoder".ST_xSystemReset )
      S_Coil( "Encoder".PH_WaitFirstMeter )
   END_RUNG
   // the same network as SCL:
   IF "Encoder".ST_xSystemReset THEN "Encoder".PH_WaitFirstMeter := TRUE; END_IF;
END_REGION

REGION Network 26: System reset done - After call buffer reset
   RUNG wire#powerrail
      Contact( "Encoder".ST_xSystemReset )
      S_Coil( "Z256_Manager".tInputData.xSystemReset )
      R_Coil( "Encoder".ST_xSystemReset )
   END_RUNG
   // the same network as SCL:
   IF "Encoder".ST_xSystemReset THEN
       "Z256_Manager".tInputData.xSystemReset := TRUE;
       "Encoder".ST_xSystemReset := FALSE;
   END_IF;
END_REGION
END_FUNCTION

FUNCTION "Z256_Output" : Void   // FC18, LAD
{ S7_Optimized_Access := 'TRUE' }
VERSION : 0.1
   VAR_TEMP
      TMP_dIndex : DInt;
      TMP_xFiring : Bool;
      TMP_xHoming : Bool;
   END_VAR
BEGIN

